// TIA Portal project "DnomaidDBMS" (V13)
// Database Management System

(* hardware
DEVICE "S71500/ET200MP station_1"  S7-1500 station
   slot 0: "Perfil soporte_0"  6ES7 590-1***0-0AA0
   slot 1: "PLC_1"  CPU 1518-4 PN/DP  6ES7 518-4AP00-0AB0  V1.8
DEVICE "HMI_1"  TP1900 Comfort
   slot 0: "HMI"  HMI  6AV2 124-0UC02-0AX0  13.0.1.0
   slot 1: "HMI_RT_1"  TP1900 Comfort  6AV2 124-0UC02-0AX0  13.0.1.0
   slot 5: "HMI_1.IE_CP_1"  Interfaz PROFINET
      slot 1: "Interfaz PROFINET_1"  Interfaz PROFINET
         slot 1: "Port_1"  Port
         slot 2: "Port_2"  Port
   slot 6: "HMI_1.IE_CP_2"  Interfaz PROFINET
      slot 1: "Interfaz PROFINET_GBit"  Interfaz PROFINET
         slot 1: "Port_1"  Port
   slot 7: "HMI_1.MPI/DP_CP_1"  Interfaz MPI/DP
*)

// ===== PLC "PLC_1"  CPU 1518-4 PN/DP =====

VAR_GLOBAL   // PLC tag table "Tabla de variables estándar"
   "System_Byte" AT %MB1 : Byte;
   "FirstScan" AT %M1.0 : Bool;
   "DiagStatusUpdate" AT %M1.1 : Bool;
   "AlwaysTRUE" AT %M1.2 : Bool;
   "AlwaysFALSE" AT %M1.3 : Bool;
   "Clock_Byte" AT %MB0 : Byte;
   "Clock_10Hz" AT %M0.0 : Bool;
   "Clock_5Hz" AT %M0.1 : Bool;
   "Clock_2.5Hz" AT %M0.2 : Bool;
   "Clock_2Hz" AT %M0.3 : Bool;
   "Clock_1.25Hz" AT %M0.4 : Bool;
   "Clock_1Hz" AT %M0.5 : Bool;
   "Clock_0.625Hz" AT %M0.6 : Bool;
   "Clock_0.5Hz" AT %M0.7 : Bool;
   "Test" AT %M10.3 : Bool;
END_VAR

TYPE "UDT_BARCODE"
AUTHOR : QLR
FAMILY : DATABASE
VERSION : 0.1
   STRUCT
      Code : "UDT_BARCODE_CODE";
      Scanner : "UDT_BARCODE_SCANNER";
   END_STRUCT;
END_TYPE

TYPE "UDT_BARCODE_CODE"
AUTHOR : QLR
FAMILY : DATABASE
VERSION : 0.1
   STRUCT
      Digit : Array[1..13] of Char;
   END_STRUCT;
END_TYPE

TYPE "UDT_BARCODE_SCANNER"
AUTHOR : QLR
FAMILY : DATABASE
VERSION : 0.1
   STRUCT
      Number : Int;
   END_STRUCT;
END_TYPE

TYPE "UDT_DATABASE_CTRL"
AUTHOR : QLR
FAMILY : DATABASE
VERSION : 0.1
   STRUCT
      FUNTION : Struct
      END_STRUCT;
      REQUEST : Struct
      END_STRUCT;
      RES01 : DInt;
   END_STRUCT;
END_TYPE

TYPE "UDT_DATABASE_DB_LIST"
VERSION : 0.1
   STRUCT
      DbNumber : Array[1..6] of Int;
      QuantityDB : Int;
   END_STRUCT;
END_TYPE

TYPE "UDT_DATABASE_M"
AUTHOR : QLR
FAMILY : DATABASE
VERSION : 0.1
   STRUCT
      RESPONSE : "UDT_DATABASE_M_RESPONSE";
      RES01 : DInt;
      REQUEST : "UDT_DATABASE_M_REQUEST";
      RES02 : DInt;
      STATUS : "UDT_DATABASE_M_STATUS";
   END_STRUCT;
END_TYPE

TYPE "UDT_DATABASE_M_REQUEST"
AUTHOR : QLR
FAMILY : DATABASE
VERSION : 0.1
   STRUCT
      Insert : Struct
      END_STRUCT;
      Query : Struct
      END_STRUCT;
      Delete : Struct
      END_STRUCT;
   END_STRUCT;
END_TYPE

TYPE "UDT_DATABASE_M_RESPONSE"
AUTHOR : QLR
FAMILY : DATABASE
VERSION : 0.1
   STRUCT
      Insert : Struct
      END_STRUCT;
      InsertData : "UDT_DATABASE_TABLE";
      Query : Struct
      END_STRUCT;
      QueryDataAvailable : "UDT_DATABASE_TABLE";
      Delete : Struct
      END_STRUCT;
      DeleteData : "UDT_DATABASE_TABLE";
   END_STRUCT;
END_TYPE

TYPE "UDT_DATABASE_M_STATUS"
AUTHOR : QLR
FAMILY : DATABASE
VERSION : 0.1
   STRUCT
      Perm : Struct
      END_STRUCT;
      Mem : Struct
      END_STRUCT;
      Fb_Fault : Bool;
      DataError : Bool;
   END_STRUCT;
END_TYPE

TYPE "UDT_DATABASE_TABLE"
AUTHOR : QLR
FAMILY : DATABASE
VERSION : 0.1
   STRUCT
      BarcodeData : "UDT_BARCODE";
      DateTime : Date_And_Time;
   END_STRUCT;
END_TYPE

TYPE "UDT_LOG"
AUTHOR : QLR
FAMILY : DATABASE
VERSION : 0.1
   STRUCT
      DatabaseTable : "UDT_DATABASE_TABLE";
      Request : Int;
   END_STRUCT;
END_TYPE

TYPE "UDT_DATABASE_DB_LIST_CONFIG"
VERSION : 0.1
   STRUCT
      DbNumber : Array[1..5] of Int;
      QuantityDB : Int;
   END_STRUCT;
END_TYPE

DATA_BLOCK "DB_GLOBAL"   // DB1
TITLE = Global
{ S7_Optimized_Access := 'FALSE' }
AUTHOR : QLR
FAMILY : dnomaiD
VERSION : 9.0
   VAR
      DataCurrentTime : Date_And_Time;
      EmptyCharDigit : Array[1..10] of Char;
      ZeroCharDigit : Array[1..10] of Char;
   END_VAR
BEGIN
END_DATA_BLOCK

DATA_BLOCK "$DB_HMI_USER"   // DB2
TITLE = DB HMI
{ S7_Optimized_Access := 'FALSE' }
AUTHOR : QLR
FAMILY : dnomaiD
VERSION : 9.0
   VAR
      GENERAL : Struct
      END_STRUCT;
      DATA_MANAGEMENT : Struct
      END_STRUCT;
      LOG : Struct
      END_STRUCT;
   END_VAR
BEGIN
END_DATA_BLOCK

DATA_BLOCK "DI_DBMS"   // DB10
TITLE = DBMS
{ S7_Optimized_Access := 'FALSE' }
AUTHOR : QLR
FAMILY : dnomaiD
VERSION : 9.0
// stored: InstanceOfName #DBMS
"#DBMS"
BEGIN
END_DATA_BLOCK

DATA_BLOCK "DB_DATABASE01"   // DB11
TITLE = Database
{ S7_Optimized_Access := 'FALSE' }
AUTHOR : QLR
FAMILY : dnomaiD
VERSION : 9.0
   VAR
      DATA : Array[1..2730] of "UDT_DATABASE_TABLE";
   END_VAR
BEGIN
END_DATA_BLOCK

DATA_BLOCK "DB_DATABASE02"   // DB12
TITLE = Database
{ S7_Optimized_Access := 'FALSE' }
AUTHOR : QLR
FAMILY : dnomaiD
VERSION : 9.0
   VAR
      DATA : Array[1..3] of "UDT_DATABASE_TABLE";
   END_VAR
BEGIN
END_DATA_BLOCK

DATA_BLOCK "DB_DATABASE03"   // DB13
TITLE = Database
{ S7_Optimized_Access := 'FALSE' }
AUTHOR : QLR
FAMILY : dnomaiD
VERSION : 9.0
   VAR
      DATA : Array[1..3] of "UDT_DATABASE_TABLE";
   END_VAR
BEGIN
END_DATA_BLOCK

DATA_BLOCK "DB_DATABASE04"   // DB14
TITLE = Database
{ S7_Optimized_Access := 'FALSE' }
AUTHOR : QLR
FAMILY : dnomaiD
VERSION : 9.0
   VAR
      DATA : Array[1..3] of "UDT_DATABASE_TABLE";
   END_VAR
BEGIN
END_DATA_BLOCK

DATA_BLOCK "DB_DATABASE05"   // DB15
TITLE = Database
{ S7_Optimized_Access := 'FALSE' }
AUTHOR : QLR
FAMILY : dnomaiD
VERSION : 9.0
   VAR
      DATA : Array[1..3] of "UDT_DATABASE_TABLE";
   END_VAR
BEGIN
END_DATA_BLOCK

DATA_BLOCK "DI_LOG"   // DB20
TITLE = Log
{ S7_Optimized_Access := 'FALSE' }
AUTHOR : QLR
FAMILY : dnomaiD
VERSION : 9.0
// stored: InstanceOfName #LOGGER
"#LOGGER"
BEGIN
END_DATA_BLOCK

DATA_BLOCK "DB_LOG"   // DB21
TITLE = Log
{ S7_Optimized_Access := 'FALSE' }
AUTHOR : QLR
FAMILY : dnomaiD
VERSION : 9.0
   VAR
      LOG : Array[1..10] of "UDT_LOG";
   END_VAR
BEGIN
END_DATA_BLOCK

DATA_BLOCK "DB_MANAGER"   // DB30
TITLE = Manager
{ S7_Optimized_Access := 'FALSE' }
AUTHOR : QLR
FAMILY : dnomaiD
VERSION : 9.0
   VAR
      LIST_DB : "UDT_DATABASE_DB_LIST_CONFIG";
      CTRL : "UDT_DATABASE_CTRL";
      DATA : "UDT_DATABASE_M";
      LOG : "UDT_LOG";
   END_VAR
BEGIN
END_DATA_BLOCK

DATA_BLOCK "CTRL_INSERT_DATA_DB"   // DB40
TITLE = Control insert data DB
{ S7_Optimized_Access := 'FALSE' }
AUTHOR : QLR
FAMILY : dnomaiD
VERSION : 9.0
// stored: InstanceOfName #CTRL_INSERT_DATA
"#CTRL_INSERT_DATA"
BEGIN
END_DATA_BLOCK

DATA_BLOCK "DB_TIMER"   // DB300
TITLE = Timer
{ S7_Optimized_Access := 'FALSE' }
AUTHOR : QLR
FAMILY : dnomaiD
VERSION : 9.0
   VAR
      TIM : Array[1..10] of IEC_TIMER;
   END_VAR
BEGIN
END_DATA_BLOCK

DATA_BLOCK "DI_SIMU_BARCODE_01"   // DB401
TITLE = Simu Barcode
{ S7_Optimized_Access := 'FALSE' }
AUTHOR : QLR
FAMILY : dnomaiD
VERSION : 9.0
// stored: InstanceOfName #SIMU_BARCODE EAN-13
"#SIMU_BARCODE EAN-13"
BEGIN
END_DATA_BLOCK

DATA_BLOCK "DI_SIMU_BARCODE_02"   // DB402
TITLE = Simu Barcode
{ S7_Optimized_Access := 'FALSE' }
AUTHOR : QLR
FAMILY : dnomaiD
VERSION : 9.0
// stored: InstanceOfName #SIMU_BARCODE EAN-13
"#SIMU_BARCODE EAN-13"
BEGIN
END_DATA_BLOCK

FUNCTION_BLOCK "#DBMS"   // FB10, STL
TITLE = DBMS
{ S7_Optimized_Access := 'FALSE' }
AUTHOR : QLR
FAMILY : dnomaiD
VERSION : 9.0
// TABLE: BarcodeData.Code | BarcodeData.Scanner | DateTime
// PRIMARY KEY: BarcodeData.Code
BEGIN

REGION Network 1: --Start--
         L     #Network_1;
         T     #P_RET_VAL.MEM;
         TAR1  #SaveAR1;
         L     STW;
         T     #SaveSTW;

         A     #Reset;
         JC    AA;
         A     #FAULT;
         S     #Status.Fb_Fault;
         JC    END;
         A     #DATA_ERROR;
         S     #Status.DataError;
         JC    AF;
   AA:   NOP   0;
         R     #FAULT;
         R     #Status.Fb_Fault;
         R     #DATA_ERROR;
         R     #Status.DataError;
   AF:   NOP   0;
END_REGION

REGION Network 2: --Timer--
         CALL  TOF , #TIME_FillAll
         ( IN := #FULL,
           PT := t#250ms,
           Q  := ,
           ET :=
         );

         A     #TIME_FillAll.Q;
         =     #Status.Mem.FillAll;
END_REGION

REGION Network 3: --Setting--
         L     #Network_3;
         T     #P_RET_VAL.MEM;
         L     #""Address_21";
         L     #""Address_9";
         XOD;
         L     8;
         /D;
         T     #LENGTH.Code;
         L     ' ';
         T     #AUX.xByte;
         CALL  FILL
         ( BVAL    := #AUX.xByte,
           RET_VAL := #P_RET_VAL.X,
           BLK     := #IniData.BarcodeData.Code
         );
         L     0;
         T     #AUX.xInt;
         L     #""Address_16";
         L     #""Address_34";
         -D;
         T     #LENGTH.PointerData;
         L     8;
         /D;
         T     #LENGTH.Data;
         CLR;
         =     #AUX.FullDatabase;
         L     5;
         T     #MaxQuantityDB;
         L     #LIST_DB.DbNumber[1];
         T     #LIST_DB_T.DbNumber[1];
         L     #LIST_DB.DbNumber[2];
         T     #LIST_DB_T.DbNumber[2];
         L     #LIST_DB.DbNumber[3];
         T     #LIST_DB_T.DbNumber[3];
         L     #LIST_DB.DbNumber[4];
         T     #LIST_DB_T.DbNumber[4];
         L     #LIST_DB.DbNumber[5];
         T     #LIST_DB_T.DbNumber[5];
         L     0;
         T     #LIST_DB_T.DbNumber[6];
         L     0;
         T     #AuxQuantityDB;

         L     #""Address_481";
         LAR1;
         L     W [ AR1 , P#0.0 ];
         T     #NDB;
         L     W [ AR1 , P#4.0 ];
         LAR1;
   bA01: NOP   0;
         OPN   DB [ #NDB ];
         L     DBW [ AR1 , P#0.0 ];
         L     0;
         ==I;
         JC    bA02;
         L     #AuxQuantityDB;
         L     1;
         +I;
         T     #AuxQuantityDB;
         L     #MaxQuantityDB;
         L     #AuxQuantityDB;
         <=I;
         JC    bA02;
         L     P#2.0;
         +AR1;
         JU    bA01;
   bA02: NOP   0;
         L     #AuxQuantityDB;
         L     1;
         <I;
         S     #FAULT;
         JC    END;
         L     #AuxQuantityDB;
         L     #MaxQuantityDB;
         >I;
         S     #FAULT;
         JC    END;
         L     #AuxQuantityDB;
         T     #QuantityDB;
         L     #QuantityDB;
         T     #LIST_DB.QuantityDB;
         T     #LIST_DB_T.QuantityDB;
END_REGION

REGION Network 4: cA..Any DB
         L     #Network_4;
         T     #P_RET_VAL.MEM;
         L     #MaxQuantityDB;
         T     #QuantityLabelDB;
         L     1;
         T     #COUNT.cA00;
         JU    cA00;
   cA00: NOP   0;
         L     #COUNT.cA00;
         JL    cAXX;
         JU    cAFF;
         JU    cA11;  //Any db[1]: First> data
         JU    cA12;  //Any db[1]: First> data, Length> all data - 1
         JU    cA13;  //Any db[1]: Last> data
         JU    cA14;  //Any db[1]: Second> data, Length> all data - 1
         JU    cA21;  //Any db[2]: First> data
         JU    cA22;  //Any db[2]: First> data, Length> all data - 1
         JU    cA23;  //Any db[2]: Last> data
         JU    cA24;  //Any db[2]: Second> data, Length> all data - 1
         JU    cA31;  //Any db[3]: First> data
         JU    cA32;  //Any db[3]: First> data, Length> all data - 1
         JU    cA33;  //Any db[3]: Last> data
         JU    cA34;  //Any db[3]: Second> data, Length> all data - 1
         JU    cA41;  //Any db[4]: First> data
         JU    cA42;  //Any db[4]: First> data, Length> all data - 1
         JU    cA43;  //Any db[4]: Last> data
         JU    cA44;  //Any db[4]: Second> data, Length> all data - 1
         JU    cA51;  //Any db[5]: First> data
         JU    cA52;  //Any db[5]: First> data, Length> all data - 1
         JU    cA53;  //Any db[5]: Last> data
         JU    cA54;  //Any db[5]: Second> data, Length> all data - 1
         JU    cA61;  //Any db[6]: First> data
         JU    cA62;  //Any db[6]: First> data, Length> all data - 1
         JU    cA63;  //Any db[6]: Last> data
         JU    cA64;  //Any db[6]: Second> data, Length> all data - 1
   cAXX: JU    cAFF;
   cA11: NOP   0;
         OPN   DB[ #LIST_DB_T.DbNumber[1]];
         L     DBNO;
         T     #PanDB[1];
         T     #PAUXnDB;  //Aux
         L     #LENGTH.Data;
         T     #AUX.LNG;  //Aux
         L     P#0.0;
         L     DW#16#84000000;
         +D;
         T     #P_ADR.I_DB[1];
         T     #P_ADR.AUX;  //Aux
         LAR1  #""Address_104";
         JU    cAFI;
   cA12: NOP   0;
         OPN   DB[ #LIST_DB_T.DbNumber[1]];
         L     DBLG;
         L     #LENGTH.Data;
         /D;
         T     #NumDataArrayDB[1];
         L     -1;
         +I;
         L     #LENGTH.Data;
         *I;
         T     #LENGTH.AllDataPushDB[1];
         T     #AUX.LNG;  //Aux
         L     #P_ADR.I_DB[1];
         T     #P_ADR.AUX;  //Aux
         LAR1  #""Address_110";
         JU    cAFI;
   cA13: NOP   0;
         L     #LENGTH.Data;
         T     #AUX.LNG;  //Aux
         OPN   DB[ #LIST_DB_T.DbNumber[1]];
         L     DBLG;
         L     #LENGTH.Data;
         -D;
         L     8;
         *D;
         L     DW#16#84000000;
         +D;
         T     #P_ADR.F_DB[1];
         T     #P_ADR.AUX;  //Aux
         LAR1  #""Address_113";
         JU    cAFI;
   cA14: NOP   0;
         L     #LENGTH.AllDataPushDB[1];
         T     #AUX.LNG;  //Aux
         L     #LENGTH.PointerData;
         L     DW#16#84000000;
         +D;
         T     #P_ADR.AUX;  //Aux
         LAR1  #""Address_115";
         JU    cAFI;
   cA21: NOP   0;
         OPN   DB[ #LIST_DB_T.DbNumber[2]];
         L     DBNO;
         T     #PanDB[2];
         T     #PAUXnDB;  //Aux
         L     #LENGTH.Data;
         T     #AUX.LNG;  //Aux
         L     P#0.0;
         L     DW#16#84000000;
         +D;
         T     #P_ADR.I_DB[2];
         T     #P_ADR.AUX;  //Aux
         LAR1  #""Address_119";
         JU    cAFI;
   cA22: NOP   0;
         OPN   DB [ #LIST_DB_T.DbNumber[2]];
         L     DBLG;
         L     #LENGTH.Data;
         /D;
         T     #NumDataArrayDB[2];
         L     -1;
         +I;
         L     #LENGTH.Data;
         *I;
         T     #LENGTH.AllDataPushDB[2];
         T     #AUX.LNG;  //Aux
         L     #P_ADR.I_DB[2];
         T     #P_ADR.AUX;  //Aux
         LAR1  #""Address_123";
         JU    cAFI;
   cA23: NOP   0;
         L     #LENGTH.Data;
         T     #AUX.LNG;  //Aux
         OPN   DB [ #LIST_DB_T.DbNumber[2]];
         L     DBLG;
         L     #LENGTH.Data;
         -D;
         L     8;
         *D;
         L     DW#16#84000000;
         +D;
         T     #P_ADR.F_DB[2];
         T     #P_ADR.AUX;  //Aux
         LAR1  #""Address_126";
         JU    cAFI;
   cA24: NOP   0;
         L     #LENGTH.AllDataPushDB[2];
         T     #AUX.LNG;  //Aux
         L     #LENGTH.PointerData;
         L     DW#16#84000000;
         +D;
         T     #P_ADR.AUX;  //Aux
         LAR1  #""Address_128";
         JU    cAFI;
   cA31: NOP   0;
         OPN   DB[ #LIST_DB_T.DbNumber[3]];
         L     DBNO;
         T     #PanDB[3];
         T     #PAUXnDB;  //Aux
         L     #LENGTH.Data;
         T     #AUX.LNG;  //Aux
         L     P#0.0;
         L     DW#16#84000000;
         +D;
         T     #P_ADR.I_DB[3];
         T     #P_ADR.AUX;  //Aux
         LAR1  #""Address_132";
         JU    cAFI;
   cA32: NOP   0;
         OPN   DB[ #LIST_DB_T.DbNumber[3]];
         L     DBLG;
         L     #LENGTH.Data;
         /D;
         T     #NumDataArrayDB[3];
         L     -1;
         +I;
         L     #LENGTH.Data;
         *I;
         T     #LENGTH.AllDataPushDB[3];
         T     #AUX.LNG;  //Aux
         L     #P_ADR.I_DB[3];
         T     #P_ADR.AUX;  //Aux
         LAR1  #""Address_136";
         JU    cAFI;
   cA33: NOP   0;
         L     #LENGTH.Data;
         T     #AUX.LNG;  //Aux
         OPN   DB[ #LIST_DB_T.DbNumber[3]];
         L     DBLG;
         L     #LENGTH.Data;
         -D;
         L     8;
         *D;
         L     DW#16#84000000;
         +D;
         T     #P_ADR.F_DB[3];
         T     #P_ADR.AUX;  //Aux
         LAR1  #""Address_139";
         JU    cAFI;
   cA34: NOP   0;
         L     #LENGTH.AllDataPushDB[3];
         T     #AUX.LNG;  //Aux
         L     #LENGTH.PointerData;
         L     DW#16#84000000;
         +D;
         T     #P_ADR.AUX;  //Aux
         LAR1  #""Address_141";
         JU    cAFI;
   cA41: NOP   0;
         OPN   DB[ #LIST_DB_T.DbNumber[4]];
         L     DBNO;
         T     #PanDB[4];
         T     #PAUXnDB;  //Aux
         L     #LENGTH.Data;
         T     #AUX.LNG;  //Aux
         L     P#0.0;
         L     DW#16#84000000;
         +D;
         T     #P_ADR.I_DB[4];
         T     #P_ADR.AUX;  //Aux
         LAR1  #""Address_145";
         JU    cAFI;
   cA42: NOP   0;
         OPN   DB[ #LIST_DB_T.DbNumber[4]];
         L     DBLG;
         L     #LENGTH.Data;
         /D;
         T     #NumDataArrayDB[4];
         L     -1;
         +I;
         L     #LENGTH.Data;
         *I;
         T     #LENGTH.AllDataPushDB[4];
         T     #AUX.LNG;  //Aux
         L     #P_ADR.I_DB[4];
         T     #P_ADR.AUX;  //Aux
         LAR1  #""Address_149";
         JU    cAFI;
   cA43: NOP   0;
         L     #LENGTH.Data;
         T     #AUX.LNG;  //Aux
         OPN   DB[ #LIST_DB_T.DbNumber[4]];
         L     DBLG;
         L     #LENGTH.Data;
         -D;
         L     8;
         *D;
         L     DW#16#84000000;
         +D;
         T     #P_ADR.F_DB[4];
         T     #P_ADR.AUX;  //Aux
         LAR1  #""Address_152";
         JU    cAFI;
   cA44: NOP   0;
         L     #LENGTH.AllDataPushDB[4];
         T     #AUX.LNG;  //Aux
         L     #LENGTH.PointerData;
         L     DW#16#84000000;
         +D;
         T     #P_ADR.AUX;  //Aux
         LAR1  #""Address_154";
         JU    cAFI;
   cA51: NOP   0;
         OPN   DB[ #LIST_DB_T.DbNumber[5]];
         L     DBNO;
         T     #PanDB[5];
         T     #PAUXnDB;  //Aux
         L     #LENGTH.Data;
         T     #AUX.LNG;  //Aux
         L     P#0.0;
         L     DW#16#84000000;
         +D;
         T     #P_ADR.I_DB[5];
         T     #P_ADR.AUX;  //Aux
         LAR1  #""Address_158";
         JU    cAFI;
   cA52: NOP   0;
         OPN   DB[ #LIST_DB_T.DbNumber[5]];
         L     DBLG;
         L     #LENGTH.Data;
         /D;
         T     #NumDataArrayDB[5];
         L     -1;
         +I;
         L     #LENGTH.Data;
         *I;
         T     #LENGTH.AllDataPushDB[5];
         T     #AUX.LNG;  //Aux
         L     #P_ADR.I_DB[5];
         T     #P_ADR.AUX;  //Aux
         LAR1  #""Address_162";
         JU    cAFI;
   cA53: NOP   0;
         L     #LENGTH.Data;
         T     #AUX.LNG;  //Aux
         OPN   DB[ #LIST_DB_T.DbNumber[5]];
         L     DBLG;
         L     #LENGTH.Data;
         -D;
         L     8;
         *D;
         L     DW#16#84000000;
         +D;
         T     #P_ADR.F_DB[5];
         T     #P_ADR.AUX;  //Aux
         LAR1  #""Address_165";
         JU    cAFI;
   cA54: NOP   0;
         L     #LENGTH.AllDataPushDB[5];
         T     #AUX.LNG;  //Aux
         L     #LENGTH.PointerData;
         L     DW#16#84000000;
         +D;
         T     #P_ADR.AUX;  //Aux
         LAR1  #""Address_167";
         JU    cAFI;
   cA61: NOP   0;
         OPN   DB[ #LIST_DB_T.DbNumber[6]];
         L     DBNO;
         T     #PanDB[6];
         T     #PAUXnDB;  //Aux
         L     #LENGTH.Data;
         T     #AUX.LNG;  //Aux
         L     P#0.0;
         L     DW#16#84000000;
         +D;
         T     #P_ADR.I_DB[6];
         T     #P_ADR.AUX;  //Aux
         LAR1  #""Address_171";
         JU    cAFI;
   cA62: NOP   0;
         OPN   DB [ #LIST_DB_T.DbNumber[6]];
         L     DBLG;
         L     #LENGTH.Data;
         /D;
         T     #NumDataArrayDB[6];
         L     -1;
         +I;
         L     #LENGTH.Data;
         *I;
         T     #LENGTH.AllDataPushDB[6];
         T     #AUX.LNG;  //Aux
         L     #P_ADR.I_DB[6];
         T     #P_ADR.AUX;  //Aux
         LAR1  #""Address_175";
         JU    cAFI;
   cA63: NOP   0;
         L     #LENGTH.Data;
         T     #AUX.LNG;  //Aux
         OPN   DB [ #LIST_DB_T.DbNumber[6]];
         L     DBLG;
         L     #LENGTH.Data;
         -D;
         L     8;
         *D;
         L     DW#16#84000000;
         +D;
         T     #P_ADR.F_DB[6];
         T     #P_ADR.AUX;  //Aux
         LAR1  #""Address_178";
         JU    cAFI;
   cA64: NOP   0;
         L     #LENGTH.AllDataPushDB[6];
         T     #AUX.LNG;  //Aux
         L     #LENGTH.PointerData;
         L     DW#16#84000000;
         +D;
         T     #P_ADR.AUX;  //Aux
         LAR1  #""Address_180";
         JU    cAFI;
   cAFI: NOP   0;
         L     B#16#10;
         T     LB[AR1, P#0.0];
         L     B#16#2;
         T     LB[AR1, P#1.0];
         L     #AUX.LNG;
         T     LW[AR1, P#2.0];
         L     #PAUXnDB;
         T     LW[AR1, P#4.0];
         L     #P_ADR.AUX;
         T     LD[AR1, P#6.0];
         L     #COUNT.cA00;
         +     1;
         T     #COUNT.cA00;
         L     #QuantityDB;
         L     #QuantityLabelDB;
         *I;
         L     #COUNT.cA00;
         <I;
         JC    cAFF;
         JU    cA00;
   //--->END
   cAFF: NOP   0;
END_REGION

REGION Network 5: cB..Status
         L     #Network_5;
         T     #P_RET_VAL.MEM;
         L     1;
         T     #COUNT.cB00;
         JU    cB00;
   cB00: NOP   0;
         L     #COUNT.cB00;
         JL    cBXX;
         JU    cBEE;  //fault
         JU    cB11;  //db[1]
         JU    cB21;  //db[2]
         JU    cB31;  //db[3]
         JU    cB41;  //db[4]
         JU    cB51;  //db[5]
         JU    cB61;  //db[6]
   cBXX: JU    cBFF;  //end
   cB11: NOP   0;
         L     #PanDB[1];
         T     #P_STATUS.nDB;
         L     #P_ADR.I_DB[1];
         T     #P_STATUS.Adr_S_DB;
         L     #P_ADR.F_DB[1];
         T     #P_STATUS.Adr_E_DB;
         JU    cBWW;
   cB21: NOP   0;
         L     #PanDB[2];
         T     #P_STATUS.nDB;
         L     #P_ADR.I_DB[2];
         T     #P_STATUS.Adr_S_DB;
         L     #P_ADR.F_DB[2];
         T     #P_STATUS.Adr_E_DB;
         JU    cBWW;
   cB31: NOP   0;
         L     #PanDB[3];
         T     #P_STATUS.nDB;
         L     #P_ADR.I_DB[3];
         T     #P_STATUS.Adr_S_DB;
         L     #P_ADR.F_DB[3];
         T     #P_STATUS.Adr_E_DB;
         JU    cBWW;
   cB41: NOP   0;
         L     #PanDB[4];
         T     #P_STATUS.nDB;
         L     #P_ADR.I_DB[4];
         T     #P_STATUS.Adr_S_DB;
         L     #P_ADR.F_DB[4];
         T     #P_STATUS.Adr_E_DB;
         JU    cBWW;
   cB51: NOP   0;
         L     #PanDB[5];
         T     #P_STATUS.nDB;
         L     #P_ADR.I_DB[5];
         T     #P_STATUS.Adr_S_DB;
         L     #P_ADR.F_DB[5];
         T     #P_STATUS.Adr_E_DB;
         JU    cBWW;
   cB61: NOP   0;
         L     #PanDB[6];
         T     #P_STATUS.nDB;
         L     #P_ADR.I_DB[6];
         T     #P_STATUS.Adr_S_DB;
         L     #P_ADR.F_DB[6];
         T     #P_STATUS.Adr_E_DB;
         JU    cBWW;
   cBEE: NOP   0;
         SET;
         S     #FAULT;
         JU    END;
   cBWW: NOP   0;
         OPN   DB[ #P_STATUS.nDB];
         LAR1  #P_STATUS.Adr_E_DB;
         L     DBB[AR1, P#0.0];
         L     ' ';
         ==I;
         =     #P_STATUS.PermInsert;
         OPN   DB[ #P_STATUS.nDB];
         LAR1  #P_STATUS.Adr_S_DB;
         L     DBB[AR1, P#0.0];
         L     ' ';
         <>I;
         =     #P_STATUS.PermOut;
         AN    #P_STATUS.PermOut;
         A     #P_STATUS.MemFull;
         =     #P_STATUS.PermPush;

         L     #COUNT.cB00;
         JL    cCXX;
         JU    cCXX;  //End
         JU    cC11;  //db[1]
         JU    cC21;  //db[2]
         JU    cC31;  //db[3]
         JU    cC41;  //db[4]
         JU    cC51;  //db[5]
         JU    cC61;  //db[6]
   cCXX: JU    cBFF;
   cC11: NOP   0;
         A     #P_STATUS.PermInsert;
         =     #Status.Perm.Insert_nDB[1];
         R     #Status.Mem.Full_nDB[1];
         A     #P_STATUS.PermOut;
         =     #Status.Perm.Out_nDB[1];
         A     #P_STATUS.PermPush;
         =     #Status.Perm.Push_nDB[1];
         JU    cCFI;
   cC21: NOP   0;
         A     #P_STATUS.PermInsert;
         =     #Status.Perm.Insert_nDB[2];
         R     #Status.Mem.Full_nDB[2];
         A     #P_STATUS.PermOut;
         =     #Status.Perm.Out_nDB[2];
         A     #P_STATUS.PermPush;
         =     #Status.Perm.Push_nDB[2];
         JU    cCFI;
   cC31: NOP   0;
         A     #P_STATUS.PermInsert;
         =     #Status.Perm.Insert_nDB[3];
         R     #Status.Mem.Full_nDB[3];
         A     #P_STATUS.PermOut;
         =     #Status.Perm.Out_nDB[3];
         A     #P_STATUS.PermPush;
         =     #Status.Perm.Push_nDB[3];
         JU    cCFI;
   cC41: NOP   0;
         A     #P_STATUS.PermInsert;
         =     #Status.Perm.Insert_nDB[4];
         R     #Status.Mem.Full_nDB[4];
         A     #P_STATUS.PermOut;
         =     #Status.Perm.Out_nDB[4];
         A     #P_STATUS.PermPush;
         =     #Status.Perm.Push_nDB[4];
         JU    cCFI;
   cC51: NOP   0;
         A     #P_STATUS.PermInsert;
         =     #Status.Perm.Insert_nDB[5];
         R     #Status.Mem.Full_nDB[5];
         A     #P_STATUS.PermOut;
         =     #Status.Perm.Out_nDB[5];
         A     #P_STATUS.PermPush;
         =     #Status.Perm.Push_nDB[5];
         JU    cCFI;
   cC61: NOP   0;
         A     #P_STATUS.PermInsert;
         =     #Status.Perm.Insert_nDB[6];
         R     #Status.Mem.Full_nDB[6];
         A     #P_STATUS.PermOut;
         =     #Status.Perm.Out_nDB[6];
         A     #P_STATUS.PermPush;
         =     #Status.Perm.Push_nDB[6];
         JU    cCFI;
   cCFI: NOP   0;
         L     #COUNT.cB00;
         +     1;
         T     #COUNT.cB00;
         L     #QuantityDB;
         >I;
         JC    cBFF;
         JU    cB00;
         JU    cBFF;
   cBFF: NOP   0;
END_REGION

REGION Network 6: cD..Move data DB_DATABASE0X<-DB_DATABASE0X+1
         L     #Network_6;
         T     #P_RET_VAL.MEM;
         L     #MaxQuantityDB;
         L     #QuantityDB;
         -I;
         L     1;
         +I;
         T     #COUNT.cD00;
         JU    cD00;
   cD00: NOP   0;
         L     #COUNT.cD00;
         JL    cDXX;
         JU    cDEE;  //fault
         JU    cD61;  //db[6]
         JU    cD51;  //db[5]
         JU    cD41;  //db[4]
         JU    cD31;  //db[3]
         JU    cD21;  //db[2]
   cDXX: JU    cDFF;  //end
   cD61: NOP   0;
         A     #Status.Perm.Out_nDB[6];
         A     #Status.Perm.Insert_nDB[5];
         JCN   cDFI;
         L     #P_RET_VAL.MEM;
         T     #P_RET_VAL.V[1];
         T     #P_RET_VAL.V[2];
         CALL  FILL
         ( BVAL    := #ANY_DB6_I,
           RET_VAL := #P_RET_VAL.V[1],
           BLK     := #ANY_DB5_F
         );
         L     #P_RET_VAL.V[1];
         L     0;
         <>I;
         S     #FAULT;
         JC    END;
         CALL  FILL
         ( BVAL    := #IniData,
           RET_VAL := #P_RET_VAL.V[2],
           BLK     := #ANY_DB6_I
         );
         L     #P_RET_VAL.V[2];
         L     0;
         <>I;
         JC    cDEE;
         R     #Status.Perm.Out_nDB[6];
         R     #Status.Perm.Insert_nDB[5];
         A     #Status.Mem.Full_nDB[6];
         S     #Status.Perm.Push_nDB[6];
         R     #Status.Mem.Full_nDB[6];
         JU    cDFF;
   cD51: NOP   0;
         A     #Status.Perm.Out_nDB[5];
         A     #Status.Perm.Insert_nDB[4];
         JCN   cDFI;
         L     #P_RET_VAL.MEM;
         T     #P_RET_VAL.V[1];
         T     #P_RET_VAL.V[2];
         CALL  FILL
         ( BVAL    := #ANY_DB5_I,
           RET_VAL := #P_RET_VAL.V[1],
           BLK     := #ANY_DB4_F
         );
         L     #P_RET_VAL.V[1];
         L     0;
         <>I;
         S     #FAULT;
         JC    END;
         CALL  FILL
         ( BVAL    := #IniData,
           RET_VAL := #P_RET_VAL.V[2],
           BLK     := #ANY_DB5_I
         );
         L     #P_RET_VAL.V[2];
         L     0;
         <>I;
         JC    cDEE;
         R     #Status.Perm.Out_nDB[5];
         R     #Status.Perm.Insert_nDB[4];
         A     #Status.Mem.Full_nDB[5];
         S     #Status.Perm.Push_nDB[5];
         R     #Status.Mem.Full_nDB[5];
         JU    cDFF;
   cD41: NOP   0;
         A     #Status.Perm.Out_nDB[4];
         A     #Status.Perm.Insert_nDB[3];
         JCN   cDFI;
         L     #P_RET_VAL.MEM;
         T     #P_RET_VAL.V[1];
         T     #P_RET_VAL.V[2];
         CALL  FILL
         ( BVAL    := #ANY_DB4_I,
           RET_VAL := #P_RET_VAL.V[1],
           BLK     := #ANY_DB3_F
         );
         L     #P_RET_VAL.V[1];
         L     0;
         <>I;
         S     #FAULT;
         JC    END;
         CALL  FILL
         ( BVAL    := #IniData,
           RET_VAL := #P_RET_VAL.V[2],
           BLK     := #ANY_DB4_I
         );
         L     #P_RET_VAL.V[2];
         L     0;
         <>I;
         JC    cDEE;
         R     #Status.Perm.Out_nDB[4];
         R     #Status.Perm.Insert_nDB[3];
         A     #Status.Mem.Full_nDB[4];
         S     #Status.Perm.Push_nDB[4];
         R     #Status.Mem.Full_nDB[4];
         JU    cDFF;
   cD31: NOP   0;
         A     #Status.Perm.Out_nDB[3];
         A     #Status.Perm.Insert_nDB[2];
         JCN   cDFI;
         L     #P_RET_VAL.MEM;
         T     #P_RET_VAL.V[1];
         T     #P_RET_VAL.V[2];
         CALL  FILL
         ( BVAL    := #ANY_DB3_I,
           RET_VAL := #P_RET_VAL.V[1],
           BLK     := #ANY_DB2_F
         );
         L     #P_RET_VAL.V[1];
         L     0;
         <>I;
         JC    cDEE;
         CALL  FILL
         ( BVAL    := #IniData,
           RET_VAL := #P_RET_VAL.V[2],
           BLK     := #ANY_DB3_I
         );
         L     #P_RET_VAL.V[2];
         L     0;
         <>I;
         JC    cDEE;
         R     #Status.Perm.Out_nDB[3];
         R     #Status.Perm.Insert_nDB[2];
         A     #Status.Mem.Full_nDB[3];
         S     #Status.Perm.Push_nDB[3];
         R     #Status.Mem.Full_nDB[3];
         JU    cDFF;
   cD21: NOP   0;
         A     #Status.Perm.Out_nDB[2];
         A     #Status.Perm.Insert_nDB[1];
         JCN   cDFI;
         L     #P_RET_VAL.MEM;
         T     #P_RET_VAL.V[1];
         T     #P_RET_VAL.V[2];
         CALL  FILL
         ( BVAL    := #ANY_DB2_I,
           RET_VAL := #P_RET_VAL.V[1],
           BLK     := #ANY_DB1_F
         );
         L     #P_RET_VAL.V[1];
         L     0;
         <>I;
         JC    cDEE;
         CALL  FILL
         ( BVAL    := #IniData,
           RET_VAL := #P_RET_VAL.V[2],
           BLK     := #ANY_DB2_I
         );
         L     #P_RET_VAL.V[2];
         L     0;
         <>I;
         JC    cDEE;
         R     #Status.Perm.Out_nDB[2];
         R     #Status.Perm.Insert_nDB[1];
         A     #Status.Mem.Full_nDB[2];
         S     #Status.Perm.Push_nDB[2];
         R     #Status.Mem.Full_nDB[2];
         JU    cDFF;
   cDEE: NOP   0;
         SET;
         S     #FAULT;
         JU    END;
   cDFI: NOP   0;
         L     #COUNT.cD00;
         +     1;
         T     #COUNT.cD00;
         JU    cD00;
         JU    cDFF;
   cDFF: NOP   0;
         JU    cE00;
   cE00: NOP   0;
         A     #Status.Mem.Full_nDB[1];
         =     #FULL;
         JCN   cEFF;
         L     #QuantityDB;
         L     1;
         >I;
         JCN   cEFF;
         A     #Status.Mem.Full_nDB[2];
         =     #FULL;
         JCN   cEFF;
         L     #QuantityDB;
         L     2;
         >I;
         JCN   cEFF;
         A     #Status.Mem.Full_nDB[3];
         =     #FULL;
         JCN   cEFF;
         L     #QuantityDB;
         L     3;
         >I;
         JCN   cEFF;
         A     #Status.Mem.Full_nDB[4];
         =     #FULL;
         L     #QuantityDB;
         L     4;
         >I;
         JCN   cEFF;
         A     #Status.Mem.Full_nDB[5];
         =     #FULL;
         L     #QuantityDB;
         L     5;
         >I;
         JCN   cEFF;
         A     #Status.Mem.Full_nDB[6];
         =     #FULL;
         JU    cEFF;
   cEFF: NOP   0;
END_REGION

REGION Network 7: cF..Data Empty auto
         JU    cF00;
   cF00: NOP   0;
         L     #Network_7;
         T     #P_RET_VAL.MEM;
         AN    #PerEmptyAuto;
         ON    #FULL;
         JC    cFFF;
         LAR1  #""Address_104";
         L     LD[AR1, P#0.0];
         T     #AUX.LD_01;
         L     LW[AR1, P#4.0];
         T     #AUX.LW_01;
         T     #PAUXnDB;
         L     LD[AR1, P#6.0];
         T     #AUX.LD_02;
         LAR1  #""Address_270";
         L     #AUX.LD_01;
         T     LD[AR1, P#0.0];
         L     #AUX.LW_01;
         T     LW[AR1, P#4.0];
         L     #AUX.LD_02;
         T     LD[AR1, P#6.0];
         OPN   DB[ #PAUXnDB];
         L     DBLG;
         L     #LENGTH.Data;
         /D;
         L     3;
         /D;
         L     1;
   cF01: NOP   0;
         T     #COUNT.cF00;
         L     #P_RET_VAL.MEM;
         T     #P_RET_VAL.V[1];
         CALL  FILL
         ( BVAL    := #IniData,
           RET_VAL := #P_RET_VAL.V[1],
           BLK     := #ANY_DB1_B
         );
         LAR1  #""Address_270";
         L     #LENGTH.PointerData;
         L     LD[AR1, P#6.0];
         +D;
         T     LD[AR1, P#6.0];
         L     #COUNT.cF00;
         LOOP  cF01;
         L     #P_RET_VAL.V[1];
         L     0;
         <>I;
         S     #FAULT;
         JC    END;
         R     #Status.Perm.Insert_nDB[1];
         A     #Status.Mem.Full_nDB[1];
         S     #Status.Perm.Push_nDB[1];
         R     #Status.Mem.Full_nDB[1];
         JU    cFFF;
   cFFF: NOP   0;
END_REGION
